// TIA Portal project "OPCServerPlanB" (V17)

(* hardware
DEVICE "S7-1500/ET200MP station_1"  S7-1500 station
   slot 0: "Rail_0"  Rack  6ES7 590-1***0-0AA0
   slot 1: "PLC_1"  CPU 1512C-1 PN  6ES7 512-1CK00-0AB0  V2.9
      slot 3: "CPU display_1"  6ES7591-1AA00-0AA0
      slot 32768: "PROFINET interface_1"  X1
         slot 32769: "Port_1"  X1 P1
         slot 32770: "Port_2"  X1 P2
      slot 34817: "Virtual CP interface port_1"  Virtual CP interface port  Virtual CP interface port
DEVICE "PC-System_1"  SIMATIC PC station
   slot 0: "SIMATIC PC station"  Rail  SIMATIC PC-Station  V1.0
      slot 125: "Stationmanager"  Station_Manager  V6.0.4
   slot 1: "HMI_RT_1"  WinCC RT Advanced  6AV2 104-0xxxx-xxxx  17.0.0.0
      slot 33792: "Computer interface"  Host interface
   slot 2: "IE general_1"  IE General  IE_CP  V8.2.0
      slot 1: "PROFINET interface"  IEGeneral.Interface.8.2.0
*)

// ===== PLC "PLC_1"  CPU 1512C-1 PN =====

VAR_GLOBAL   // PLC tag table "Default tag table"
   "System_Byte" AT %MB1 : Byte;
   "FirstScan" AT %M1.0 : Bool;
   "DiagStatusUpdate" AT %M1.1 : Bool;
   "AlwaysTRUE" AT %M1.2 : Bool;
   "AlwaysFALSE" AT %M1.3 : Bool;
   "Clock_Byte" AT %MB0 : Byte;
   "Clock_10Hz" AT %M0.0 : Bool;
   "Clock_5Hz" AT %M0.1 : Bool;
   "Clock_2.5Hz" AT %M0.2 : Bool;
   "Clock_2Hz" AT %M0.3 : Bool;
   "Clock_1.25Hz" AT %M0.4 : Bool;
   "Clock_1Hz" AT %M0.5 : Bool;
   "Clock_0.625Hz" AT %M0.6 : Bool;
   "Clock_0.5Hz" AT %M0.7 : Bool;
END_VAR

DATA_BLOCK "DATA_OPC"   // DB1
{ S7_Optimized_Access := 'TRUE' }
VERSION : 0.1
   VAR
      "Cart_storage_1.n_carts" : DInt;
      "Cart_storage_1.start.signal" : LReal;
      "Cart_storage_1.v_carros" : LReal;
      "Unit_Sterilizer_1.st1.batch_in_ster.signal" : LReal;
      "Unit_Sterilizer_1.st1.batch_ready.signal" : LReal;
      "Unit_Sterilizer_1.st1.TR" : LReal;
      "Unit_Sterilizer_1.v_st1.Ap.signal" : LReal;
   END_VAR
   VAR RETAIN
      "Unit_Sterilizer_1.stage.signal" : LReal;
   END_VAR
   VAR
      "TIME" : LReal;
   END_VAR
BEGIN
END_DATA_BLOCK

DATA_BLOCK "DATA_PID"   // DB2
{ S7_Optimized_Access := 'TRUE' }
VERSION : 0.1
   VAR
      "Unit_Sterilizer_1.slpr" : LReal;
      "Unit_Sterilizer_1.st1.Trm" : LReal;
      ramp_enable : Bool;
      "Unit_Sterilizer_1.st1.Trm_out_delayed" : LReal;
      range_pv_min : LReal;
      range_pv_max : LReal;
      range_pv_min_scaled : LReal;
      range_pv_max_scaled : LReal;
      pv_min_scaled : LReal;
      pv_max_scaled : LReal;
      "Unit_Sterilizer_1.st1.TR_scaled" : LReal;
      "Unit_Sterilizer_1.st1.Trm_out_scaled" : LReal;
      track_mode : Bool;
      active_pos : LReal;
      Timer_enable : Bool;
      "Timer" : Time;
      "Unit_Sterilizer_1.st1.Trm_out_substitute" : LReal;
      Enable_Stage_2 : Bool;
      Enable_STOP : Bool;
   END_VAR
BEGIN
END_DATA_BLOCK

// folder: System blocks/Program resources

DATA_BLOCK "IEC_Timer_0_DB"   // DB3
{ S7_Optimized_Access := 'TRUE' }
AUTHOR : Simatic
FAMILY : IEC
NAME : IEC_TMR
VERSION : 1.0
// stored: InstanceOfName IEC_TIMER
"IEC_TIMER"
BEGIN
END_DATA_BLOCK

// folder: (top level)

FUNCTION "FCN_LOGIC" : Void   // FC1, SCL
{ S7_Optimized_Access := 'TRUE' }
VERSION : 0.1
BEGIN
   // HABILITAR CARGA DE CARROS
   IF LREAL_TO_INT("DATA_OPC"."Unit_Sterilizer_1.stage.signal") = 0 THEN
       "DATA_PID".track_mode := TRUE;
       "DATA_PID".ramp_enable := TRUE;
   END_IF;

   //HABILITAR CALENTAMIENTO
   IF LREAL_TO_INT("DATA_OPC"."Cart_storage_1.start.signal") = 1 THEN
       IF LREAL_TO_INT("DATA_OPC"."Unit_Sterilizer_1.st1.batch_ready.signal") = 1 THEN
           "DATA_OPC"."Unit_Sterilizer_1.stage.signal" := 1.0;
       END_IF;
   END_IF;


   //ETAPA CALENTAMIENTO - RAMPA
   IF LREAL_TO_INT("DATA_OPC"."Cart_storage_1.start.signal") = 1 THEN
           IF LREAL_TO_INT("DATA_OPC"."Unit_Sterilizer_1.stage.signal") = 1 THEN
               IF LREAL_TO_INT("DATA_OPC"."Unit_Sterilizer_1.st1.batch_ready.signal") = 1 THEN
                   "DATA_PID".track_mode := FALSE;
                   "DATA_PID".ramp_enable := FALSE;
               END_IF;
           END_IF;
   END_IF;

   // ETAPA CALENTAMIENTO - MANTENIMIENTO
   IF LREAL_TO_INT("DATA_OPC"."Cart_storage_1.start.signal") = 1 THEN
       IF LREAL_TO_INT("DATA_OPC"."Unit_Sterilizer_1.stage.signal") = 1 THEN
           IF "SP-PID".UpperLimit_Active = TRUE THEN
               "DATA_PID".Timer_enable := TRUE;
           END_IF;
       END_IF;
   END_IF;

   IF "DATA_PID".Timer_enable = TRUE THEN
       "DATA_PID".Timer := T#1420000ms;
       "IEC_Timer_0_DB".TON(IN := "DATA_PID".Timer_enable,
                            PT := "DATA_PID".Timer,
                            Q => "DATA_PID".Enable_Stage_2);
       "DATA_PID".Timer_enable := FALSE;
   END_IF;

   IF "DATA_PID".Enable_Stage_2 = TRUE THEN
       "DATA_OPC"."Unit_Sterilizer_1.stage.signal" := 2.0;
       "DATA_PID".track_mode := TRUE;
       "DATA_PID".ramp_enable := TRUE;
   END_IF;

   //ETAPA ENFRIAMIENTO
   IF LREAL_TO_INT("DATA_OPC"."Unit_Sterilizer_1.stage.signal") = 2 THEN
       "DATA_PID".track_mode := TRUE;
       "DATA_PID".track_mode := TRUE;
       "DATA_PID".active_pos := 0.0;
       IF LREAL_TO_INT("DATA_OPC"."Unit_Sterilizer_1.st1.TR") < 320 THEN
            "DATA_OPC"."Cart_storage_1.start.signal" := 0.0;
            "DATA_OPC"."Unit_Sterilizer_1.stage.signal" := 0.0;
       END_IF;
   END_IF;

   //SETEO A CEROS DE VALORES DE PROCESO
   IF "DATA_PID".Enable_STOP = TRUE THEN
       "DATA_OPC"."Cart_storage_1.start.signal" := 0.0;
       "DATA_OPC"."Unit_Sterilizer_1.stage.signal" := 0.0;
       "DATA_OPC"."Cart_storage_1.v_carros" := 0.0;
       "DATA_OPC"."Unit_Sterilizer_1.v_st1.Ap.signal" := 0.0;
       ;
   END_IF;
END_FUNCTION

ORGANIZATION_BLOCK "Main"   // OB1, SCL, ProgramCycle
TITLE = "Main Program Sweep (Cycle)"
{ S7_Optimized_Access := 'TRUE' }
VERSION : 0.1
   VAR_INPUT
      Initial_Call : Bool;   // Initial call of this OB
      Remanence : Bool;   // =True, if remanent data are available
   END_VAR
BEGIN
   "FCN_LOGIC"();
END_ORGANIZATION_BLOCK

ORGANIZATION_BLOCK "PID Cyclic interrupt"   // OB30, LAD, CyclicInterrupt
{ S7_Optimized_Access := 'TRUE' }
VERSION : 0.1
   VAR_INPUT
      Initial_Call : Bool;   // Initial call of this OB
      Event_Count : Int;   // Events discarded
   END_VAR
   VAR_TEMP
      error_1 : Bool;
      error_2 : Bool;
      status_1 : Word;
      status_2 : Word;
   END_VAR
   VAR_TEMP   // added for the SCL form of the ladder/FBD networks
      _w1 : Bool;
   END_VAR
BEGIN

REGION Network 1
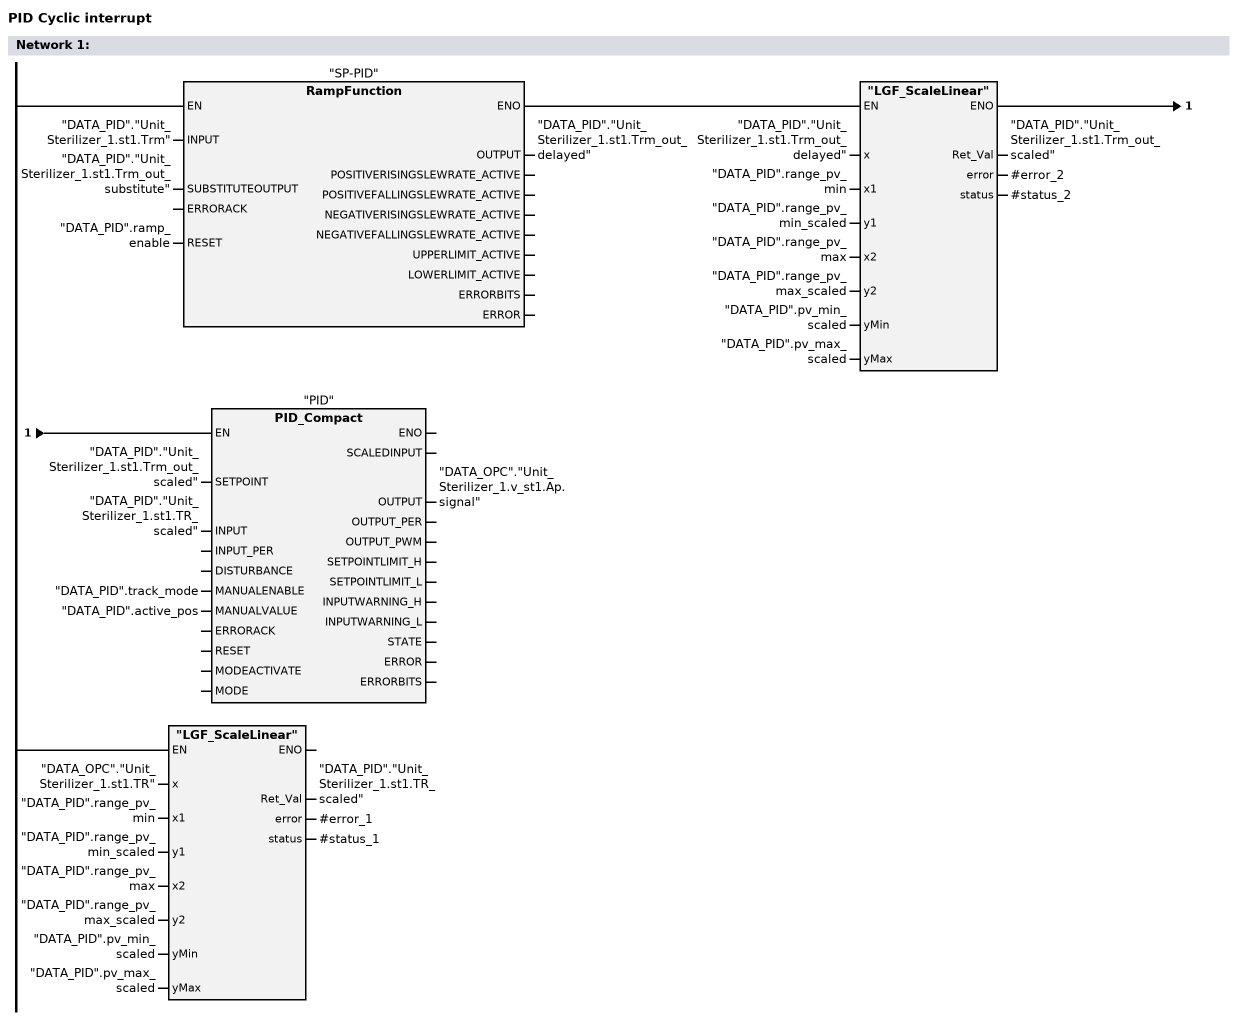
   // ENO of a box is taken as its EN; it also drops when the box reports an error
   "SP-PID"(Input := "DATA_PID"."Unit_Sterilizer_1.st1.Trm",   // RampFunction
            SubstituteOutput := "DATA_PID"."Unit_Sterilizer_1.st1.Trm_out_substitute",
            Reset := "DATA_PID".ramp_enable,
            Output => "DATA_PID"."Unit_Sterilizer_1.st1.Trm_out_delayed");
   "DATA_PID"."Unit_Sterilizer_1.st1.Trm_out_scaled" := "LGF_ScaleLinear"(x := "DATA_PID"."Unit_Sterilizer_1.st1.Trm_out_delayed",
                           x1 := "DATA_PID".range_pv_min,
                           y1 := "DATA_PID".range_pv_min_scaled,
                           x2 := "DATA_PID".range_pv_max,
                           y2 := "DATA_PID".range_pv_max_scaled,
                           yMin := "DATA_PID".pv_min_scaled,
                           yMax := "DATA_PID".pv_max_scaled,
                           error => #error_2,
                           status => #status_2,
                           ENO => #_w1);
   IF #_w1 THEN
       "PID"(Setpoint := "DATA_PID"."Unit_Sterilizer_1.st1.Trm_out_scaled",   // PID_Compact
             Input := "DATA_PID"."Unit_Sterilizer_1.st1.TR_scaled",
             ManualEnable := "DATA_PID".track_mode,
             ManualValue := "DATA_PID".active_pos,
             Output => "DATA_OPC"."Unit_Sterilizer_1.v_st1.Ap.signal");
   END_IF;
   "DATA_PID"."Unit_Sterilizer_1.st1.TR_scaled" := "LGF_ScaleLinear"(x := "DATA_OPC"."Unit_Sterilizer_1.st1.TR",
                           x1 := "DATA_PID".range_pv_min,
                           y1 := "DATA_PID".range_pv_min_scaled,
                           x2 := "DATA_PID".range_pv_max,
                           y2 := "DATA_PID".range_pv_max_scaled,
                           yMin := "DATA_PID".pv_min_scaled,
                           yMax := "DATA_PID".pv_max_scaled,
                           error => #error_1,
                           status => #status_1);
END_REGION
END_ORGANIZATION_BLOCK

ORGANIZATION_BLOCK "RampReset Cyclic interrupt"   // OB31, SCL, CyclicInterrupt
{ S7_Optimized_Access := 'TRUE' }
VERSION : 0.1
   VAR_INPUT
      Initial_Call : Bool;   // Initial call of this OB
      Event_Count : Int;   // Events discarded
   END_VAR
BEGIN
   IF "DATA_OPC"."Unit_Sterilizer_1.stage.signal" = 1 THEN
       IF "DATA_PID".ramp_enable = TRUE THEN
           "SP-PID".Reset := TRUE;
           "DATA_PID".ramp_enable := FALSE;
       ELSE
           "SP-PID".Reset := FALSE;
       END_IF;
   END_IF;
END_ORGANIZATION_BLOCK

ORGANIZATION_BLOCK "Startup"   // OB100, SCL, Startup
TITLE = "Complete Restart"
{ S7_Optimized_Access := 'TRUE' }
VERSION : 0.1
   VAR_INPUT
      LostRetentive : Bool;   // True if retentive data are lost
      LostRTC : Bool;   // True if date and time are lost
   END_VAR
BEGIN
   // Inicialización
   // PID
   "DATA_PID"."Unit_Sterilizer_1.st1.Trm" := 394.5;
   "DATA_PID"."Unit_Sterilizer_1.st1.Trm_out_substitute" := 328.0;
   "DATA_PID"."Unit_Sterilizer_1.slpr" := 0.028;
   "DATA_PID".range_pv_min := 300;
   "DATA_PID".range_pv_max := 400;
   "DATA_PID".range_pv_min_scaled := 0.0;
   "DATA_PID".range_pv_max_scaled := 100.0;
   "DATA_PID".pv_min_scaled := 0.0;
   "DATA_PID".pv_max_scaled := 100.0;
   "DATA_PID".active_pos := 0;

   //RAMPA
   "SP-PID".PositiveRisingSlewRate := 0.028;
   "SP-PID".UpperLimit := LREAL_TO_REAL("DATA_PID"."Unit_Sterilizer_1.st1.Trm");
   "DATA_PID".ramp_enable := TRUE;

   //TEMPORIZADOR
   "DATA_PID".Timer_enable := FALSE;

   //PROCESO
   "DATA_OPC"."Cart_storage_1.v_carros" := 0.0;
   "DATA_OPC"."Unit_Sterilizer_1.stage.signal" := 0.0;
   "DATA_OPC"."Cart_storage_1.start.signal" := 0.0;
   "DATA_PID".Enable_STOP := FALSE;
   "DATA_OPC"."Unit_Sterilizer_1.v_st1.Ap.signal" := 0.0;

   //PID PARAMETERS DISABLED
   "PID".CycleTime.EnEstimation := FALSE;
   "PID".CycleTime.EnMonitoring := FALSE;
END_ORGANIZATION_BLOCK

// folder: LGF/04 Math operations

FUNCTION "LGF_ScaleLinear" : LReal   // FC10039, SCL
TITLE = LGF_ScaleLinear
{ S7_Optimized_Access := 'TRUE' }
AUTHOR : Siemens_Digital_Industry_Support
FAMILY : LGF
NAME : LGF_ScaleLinear
// This function scales an input variable (`LReal`) via a linear straight-line equation. / Diese Funktion skaliert eine Eingangsgröße (`LReal`) über eine lineare Geradengleichung.
   VAR_INPUT
      x : LReal;   // Input value `x` to be scaled. / Eingangswert `x` der skaliert werden soll.
      x1 : LReal;   // Point 1 (P1) -`x` coordinate of the linear function. / Punkt 1 (P1) - `x` Koordinate der linearen Funktion.
      y1 : LReal;   // Point 1 (P1) -`y` coordinate of the linear function. / Punkt 1 (P1) - `y` Koordinate der linearen Funktion.
      x2 : LReal;   // Point 2 (P2) -`x` coordinate of the linear function. / Punkt 2 (P2) - `x` Koordinate der linearen Funktion.
      y2 : LReal;   // Point 2 (P2) -`y` coordinate of the linear function. / Punkt 2 (P2) - `y` Koordinate der linearen Funktion.
      yMin : LReal;   // Lower limit value of the output. / Unterer Grenzwert des Ausgangs.
      yMax : LReal;   // High limit value of the output. / Oberer Grenzwert des Ausgangs.
   END_VAR
   VAR_OUTPUT
      error : Bool;   // FALSE: No error TRUE: An error occurred during the execution of the FB / FALSE: Kein Fehler TRUE: Während der Ausführung des FB ist ein Fehler aufgetreten
      status : Word;   // 16#0000-16#7FFF: Status of the FB 16#8000-16#FFFF: Error identification (see following Table) / 16#0000-16#7FFF: Status des FB 16#8000-16#FFFF: Fehleridentifikation (siehe folgende Tabelle)
   END_VAR
   VAR_TEMP
      tempY : LReal;   // Temp scaled value `y` / Temp Skalierter Wert `y`
      tempStatus : Word;   // Temp status memory / Temp Status Variable
   END_VAR
   // Ret_Val : Scaled output value `y` / Skalierter Ausgangswert `y`
   VAR CONSTANT
      STATUS_FINISHED_NO_ERROR : Word := 16#0000;   // Status: Execution finished without errors. / Status: Abarbeitung ohne Fehler beendet
      ERR_LOW_LIM_OVER_UP_LIM : Word := 16#8200;   // Error: Lower limit value `yMin` is greater than high limit value `yMax`. / Fehler: Unterer Grenzwert `yMin` ist größer als oberer Grenzwert `yMax`.
      WARN_Y_LIMITED_TO_YMIN : Word := 16#6001;   // Warning: Output value limited to `yMin` / Warnung: Ausgabewert auf `yMin` begrenzt
      WARN_Y_LIMITED_TO_YMAX : Word := 16#6002;   // Warning: Output value limited to `yMax` / Warnung: Ausgabewert auf `yMax` begrenzt
      PRECISION : LReal := 1.0E-06;   // Accuracy with which the two numbers are considered equal / Genauigkeit mit welcher die beiden Werte vergleichen werden und auf "Gleichheit" geprüft werden
   END_VAR
BEGIN
   REGION BLOCK INFO HEADER
     //===============================================================================
     // SIEMENS AG / (c)Copyright 2017
     //-------------------------------------------------------------------------------
     // Title:            LGF_ScaleLinear
     // Comment/Function: This function scales an input variable (`LReal`) via a linear straight-line equation.
     // Library/Family:   LGF(Library General Functions)
     // Author:           Siemens Digital Industry Support
     // Tested with:      S7-PLCSIM Advanced V2.0 SP1
     // Engineering:      TIA Portal V14 Upd 1
     // Restrictions:     ENO mechanism is not used, Error handling done by error and status
     // Requirements:     PLC (S7-1200 / S7-1500)
     //-------------------------------------------------------------------------------
     // Change log table:
     // Version  | Date       | Expert in charge       | Changes applied
     //----------|------------|------------------------|------------------------------
     // 01.00.00 | 27.01.2017 | Siemens Industry Online Support
     //                         First released version
     // 01.00.01 | 17.08.2018 | Siemens Industry Online Support
     //                         Upgrade: TIA V15 Update 2
     // 01.00.02 | 23.11.2018 | Siemens Industry Online Support
     //                         Upgrade: TIA V15.1
     // 02.00.00 | 25.01.2019 | Simatic Systems Support
     //                         Data type changed from Variant to LReal
     // 02.00.01 | 25.06.2019 | Simatic Systems Support
     //                         Standard header and block parameters update, status parameter added
     //                         LReal value comparison added
     //                         Result parameter changed to return value of FC for use in SCL
     //                         Warning number changed to range of 16#6xxx
     //                         refactor variable handling and extract returns in between the code
     //                         add ENO handling
     // 03.00.00 | 23.04.2020 | Simatic Systems Support | Set version to V3.0.0
     //                         harmonize the version of the whole library
     // 03.00.01 | 12.11.2020 | Simatic Systems Support
     //                         Insert documentation
     //                         Move to folder "Math operations"
     //=============================================================================
   END_REGION Block info header

   REGION DESCRIPTION
     (/*The function linearly scales an input variable (e.g. an analog input value) to a specific output variable (e.g. level).

   To determine the output variable, the following linear equation is used in the function:

   $$
    x = \frac{y_2 - y_1}{x_2 - x_1} * (x - x_1) + y_1
   $$

   The straight line is described by the two points, P1 and P2. You specify the points as a Cartesian coordinate system using x and y coordinates.

   Note
   :    If the values of the parameters `x1` and `x2` are the same, the value of `y1` is output on output `y`.

   ---

   By specifying `yMin` and `yMax` you can restrict the calculated value of `y` to a range limited at top and bottom. Thus, you avoid override and underride ranges.

   Figure: Graphical representation

   ![LGF_ScaleLinear - Principle of operation](LGF_ScaleLinear.PNG "LGF_ScaleLinear - Principle of operation")

   #### Example

   A signal from 4 to 20mA is applied on an analog input module. This signal is converted to the CPU internal value from 0 to 27648 to measure a level. 0 corresponds to a level of 0.0m and 27648 to a level of 1.7m.

   The block must then be parameterized as follows:  
   * P2: $x1 = 0$; $y1 = 0.0$
   * P2: $x2 = +27648$; $y2 = 1.7$
   * $yMin = 0.0$; $yMax = 1.7$;
   Die Funktion skaliert eine Eingangsgröße (z. B. ein Analogeingangswert) linear auf eine bestimmte Ausgangsgröße (z. B. Füllstand).

   Zur Bestimmung der Ausgangsgröße wird in der Funktion folgende lineare Geradengleichung angewendet:

   $$
    x = \frac{y_2 - y_1}{x_2 - x_1} * (x - x_1) + y_1
   $$

   Die Gerade wird durch die zwei Punkte, P1 und P2, beschrieben. Die Punkte geben Sie im Sinne eines kartesischen Koordinatensystems durch x- und y-Koordinaten vor.

   Hinweis
   :    Falls die Werte der Parameter `x1` und `x2` gleich sind, wird am Ausgang `y` der Wert von `y1` ausgegeben.

   ---

   Mit der Angabe von `yMin` und `yMax` können Sie den berechneten Wert von `y` auf einen unten und oben begrenzten Bereich einschränken. Somit vermeiden Sie Über- und Untersteuerungsbereiche.

   Abbildung: Graphische Darstellung

   ![LGF_ScaleLinear - Funktionsweise](LGF_ScaleLinear.PNG "LGF_ScaleLinear - Funktionsweise")

   #### Beispiel

   An einer Analogeingangsbaugruppe liegt ein Signal von 4 bis 20mA an. Dieses Signal wird zu dem CPU-internen Wert von 0 bis 27648 gewandelt, um einen Füllstand zu messen. Dabei entsprechen 0 dem Füllstand 0,0m und 27648 dem Füllstand 1,7m.

   Den Baustein müssen Sie dann wie folgt parametrieren:  
   * P2: $x1 = 0$; $y1 = 0,0$
   * P2: $x2 = +27648$; $y2 = 1,7$
   * $yMin = 0,0$; $yMax = 1,7$;*/)
   END_REGION DESCRIPTION

   REGION INITIALISATION
     #tempY := 0.0;
     #tempStatus := #STATUS_FINISHED_NO_ERROR;
   END_REGION

   REGION CONVERT
     // check if limits in a plausible range
     // --> higher limit has to be greater than lower limit
     IF (#yMin > #yMax) THEN
       #tempY := 0.0;
       #tempStatus := #ERR_LOW_LIM_OVER_UP_LIM;

     ELSE// no error, process scaling
       // Scale algorithm
       IF (ABS(#x1 - #x2) <= (#PRECISION * ABS(#x1))) THEN
         //The slope is approximately ZERO.
         //Special CASE, use a different equation, NOT "y = m*x+t", instead you use "x = y1"
         #tempY := #y1;
       ELSE
         // resolved equation --> F(x) = y = m*x+t, where m = slope/gradient, t = intercept
         #tempY := (#y2 - #y1) / (#x2 - #x1) * (#x - #x1) + #y1;
       END_IF;

       // Check if upper or lower limit is exceeded
       IF (#tempY < #yMin) THEN
         #tempY := #yMin;
         #tempStatus := #WARN_Y_LIMITED_TO_YMIN;  // set warning indicator
       ELSIF (#tempY > #yMax) THEN
         #tempY := #yMax;
         #tempStatus := #WARN_Y_LIMITED_TO_YMAX;  // set warning indicator
       END_IF;
     END_IF;
   END_REGION

   REGION OUTPUTS  
     // set status and error output
     #status := #tempStatus;
     #error := #tempStatus.%X15;
     // set return value
     #LGF_ScaleLinear := #tempY;
     //ENO mechanism is not used - forced to true.
     ENO := TRUE;
   END_REGION
END_FUNCTION

(* ===== HMI "HMI_RT_1" =====
system functions are stored by id; their names below are inferred from use
connection "HMI_Connection_2": ETHERNET, S7_1500_OMS

HMI tags "Default tag table"
   "HMI_Tag_Cart_storage_1.cart_in" : DInt = PLC DATA_OPC."Cart_storage_1.n_carts" AT %DB1.DBW0, 1 s
   "HMI_Tag_Cart_storage_1.start.signal" : LReal = PLC DATA_OPC."Cart_storage_1.start.signal" AT %DB1.DBD0, 1 s
   "HMI_Tag_Cart_storage_1.v_carros" : LReal = PLC DATA_OPC."Cart_storage_1.v_carros" AT %DB1.DBX0.0, 1 s
   "HMI_Tag_Unit_Sterilizer_1.st1.batch_in_ster.signal" : LReal = PLC DATA_OPC."Unit_Sterilizer_1.st1.batch_in_ster.signal" AT %DB1.DBX0.0, 1 s
   "HMI_Tag_Unit_Sterilizer_1.st1.batch_ready.signal" : LReal = PLC DATA_OPC."Unit_Sterilizer_1.st1.batch_ready.signal" AT %DB1.DBX0.0, 1 s
   "HMI_Tag_Unit_Sterilizer_1.st1.TR" : LReal = PLC DATA_OPC."Unit_Sterilizer_1.st1.TR" AT %DB1.DBX0.0, 1 s
   "HMI_Tag_Unit_Sterilizer_1.v_st1.Ap.signal" : LReal = PLC DATA_OPC."Unit_Sterilizer_1.v_st1.Ap.signal" AT %DB1.DBX0.0, 1 s
   "HMI_Tag_Unit_Sterilizer_1.stage.signal" : LReal = PLC DATA_OPC."Unit_Sterilizer_1.stage.signal" AT %DB1.DBX0.0, 1 s
   "HMI_Tag_TIME" : LReal = PLC DATA_OPC.TIME AT %DB1.DBX0.0, 1 s
   "HMI_Tag_Unit_Sterilizer_1.st1.Trm" : LReal = PLC DATA_PID."Unit_Sterilizer_1.st1.Trm" AT %DB1.DBX0.0, 1 s
   "HMI_Tag_Unit_Sterilizer_1.st1.Trm_out_delayed" : LReal = PLC DATA_PID."Unit_Sterilizer_1.st1.Trm_out_delayed" AT %DB1.DBX0.0, 1 s

text list "VALVE_ON_OFF": 0 'CERRADA'; 1 'CERRADA'; 2 'ABIERTA'

text list "ESTADO DE CARGA": 0 'CARGANDO'; 1 'LISTO'

text list "VELOCIDAD": 20 '20'; 10 '10'; 0 '0'; 30 '30'; 40 '40'; 50 '50'; 60 '60'; 70 '70'; 80 '80'; 90 '90'; 100 '100'; 110 '110'; 120 '120'; 130 '130'; 140 '140'; 150 '150'; 160 '160'; 170 '170'; 180 '180'; 190 '190'; 200 '200'

screen "COVER" 1920x1200
   TextField "Text field_1" at 0,213 size 1911x56; Text 'UN ENTORNO VIRTUAL CON CONTROLADORES LÓGICOS PROGRAMABLES (PLC):'
   TextField "Text field_2" at 0,265 size 1913x58; Text 'APLICACIÓN EN EVALUACIÓN DE ESTRATEGIAS DE CONTROL'
   Button "Button_1" at 836,532 size 212x76; TextOff 'INICIAR'
      on Click: ActivateScreen("HOME", 0)
   GraphicView "Graphic view_1" at 68,652 size 534x320; Picture "logouva-removebg-preview"
   GraphicView "Graphic view_2" at 678,652 size 600x356; Picture "logoisp-removebg-preview"
   GraphicView "Graphic view_3" at 1416,672 size 400x300; Picture "logo_cspuva"
   Button "Button_2" at 1676,1096 size 212x76; TextOff 'SALIR'
      on Click: StopRuntime(0)

Template "HOME" 1920x1200
   TextField "Template_Text field_1" at 1424,16 size 467x68; Text 'ESTADO DE LA CPU-PLC'
   Button "Button_2" at 1676,1096 size 212x76; TextOff 'SALIR'
      on Click: StopRuntime(0)
   Button "Button_1" at 1464,91 size 184x60; TextOff 'INICIAR'
      on Click: function_f249594b("HMI_Connection_2", 8)
   Button "Button_3" at 1678,92 size 184x58; TextOff 'DETENER'
      on Click: function_f249594b("HMI_Connection_2", 4)
   TextField "Template_Text field_2" at 39,16 size 1187x68; Text 'UNIDAD DE PROCESO DE ESTERILIZACIÓN'
   TextField "Template_Text field_3" at 1422,204 size 482x68; Text 'PROCESO POR LOTES'
   Button "Button_4" at 1464,260 size 184x60; TextOff 'INICIAR'
      on Click: SetTag("HMI_Tag_Cart_storage_1.start.signal", 1)
      on Activate: SetTag("HMI_Tag_Cart_storage_1.start.signal", 1)
   Button "Button_5" at 1680,262 size 184x58; TextOff 'DETENER'
      on Click: SetTag("HMI_Tag_Cart_storage_1.start.signal", 0)
   IOField "Template_I/O field_1" at 1464,347 size 62x59; FormatPattern 9
      ProcessValue <- "HMI_Tag_Unit_Sterilizer_1.stage.signal"
   TextField "Template_Text field_4" at 1545,323 size 345x68; Text '0 - CARGA'
   TextField "Template_Text field_5" at 1546,356 size 343x68; Text '1 - CALENTAMIENTO'
   TextField "Template_Text field_6" at 1546,389 size 344x68; Text '2 - ENFRIAMIENTO'

screen "HOME" 1920x1200, template "HOME"
   GraphicView "Graphic view_1" at 3,103 size 1246x964; Picture "HMI_5"
   IOField "I/O field_2" at 535,236 size 88x32; FormatPattern 999; Unit  %
      ProcessValue <- "HMI_Tag_Unit_Sterilizer_1.v_st1.Ap.signal"
   IOField "I/O field_3" at 1132,1067 size 205x32; FormatPattern 99
      ProcessValue <- "HMI_Tag_Cart_storage_1.cart_in"
   TextField "Text field_1" at 792,1068 size 209x32; Text 'NRO DE CARROS'
   TextField "Text field_2" at 792,1097 size 337x34; Text 'VELOCIDAD [CARROS/H]'
   IOField "I/O field_6" at 966,281 size 123x32; FormatPattern 999; Unit  K
      ProcessValue <- "HMI_Tag_Unit_Sterilizer_1.st1.TR"
   TextField "Text field_3" at 863,227 size 117x29; Text 'SP'
   TextField "Text field_4" at 863,282 size 108x30; Text 'PV'
   IOField "I/O field_7" at 966,253 size 123x32; FormatPattern 999; Unit  K
      ProcessValue <- "HMI_Tag_Unit_Sterilizer_1.st1.Trm_out_delayed"
   TextField "Text field_5" at 863,254 size 116x29; Text 'SP OUT'
   TextField "Text field_6" at 1295,472 size 603x50; Text 'TENDENCIAS'
   SymbolicIOField "Symbolic I/O field_1" at 626,388 size 199x32; TextOff '0'; TextOn '1'; TextList "VALVE_ON_OFF"
      ProcessValue <- "HMI_Tag_Unit_Sterilizer_1.stage.signal"
   TrendView "Trend view_1" at 1297,565 size 600x208
   TextField "Text field_8" at 792,1124 size 243x34; Text 'CARROS/LOTE : 12'
   IOField "I/O field_1" at 966,224 size 123x32; FormatPattern 999; Unit  K
      ProcessValue <- "HMI_Tag_Unit_Sterilizer_1.st1.Trm"
   SymbolicIOField "Symbolic I/O field_2" at 1132,1096 size 205x32; TextOff '0'; TextOn '1'; TextList "VELOCIDAD"
      ProcessValue <- "HMI_Tag_Cart_storage_1.v_carros"
   TextField "Text field_9" at 1294,514 size 603x50; Text 'TT-01'
   TextField "Text field_10" at 1295,795 size 603x50; Text 'TV-01'
   TrendView "Trend view_2" at 1298,844 size 600x208
*)